   "DB_SDC_GLOBAL_EMS_ID_ACT" : Int = PLC DB_SDC_GLOBAL.EMS_ID_ACT AT %DB3700.DBW0, 1 s   // Aktuelle Anzahl der EMS-Treiber / Current quantity of EMS drivers
   "DB_SDC_GLOBAL_SYNCH[3].MAX_FAKT" : Real = PLC DB_SDC_GLOBAL.SYNCH[3].MAX_FAKT AT %DB3700.DBD214, 1 s   // Faktor für maximale Synchronisiergeschwindigkeit / Faktor Speed for Synchron MAX
   "DB_SDC_GLOBAL_SYNCH[13].SET_DIST" : Int = PLC DB_SDC_GLOBAL.SYNCH[13].SET_DIST AT %DB3700.DBW384, 1 s   // Set point value: distance (mm)
   "DB_SDC_GLOBAL_LIMITS[3].RAPID_SLOW" : Int = PLC DB_SDC_GLOBAL.LIMITS[3].RAPID_SLOW AT %DB3700.DBW518, 1 s   // Umstellung Begrenzung auf Abstand (mm), Einschränkung / Changeover limit of distance (mm), limitation
   "DB_SDC_GLOBAL_SYNCH[3].K" : Real = PLC DB_SDC_GLOBAL.SYNCH[3].K AT %DB3700.DBD210, 1 s   // erreichen von Synchron Faktor / gain for Synchron Faktor
   "DB_SDC_GLOBAL_SYNCH[13].SYNCH_DIST" : Int = PLC DB_SDC_GLOBAL.SYNCH[13].SYNCH_DIST AT %DB3700.DBW386, 1 s   // Start synchron distance value: distance (mm)
   "DB_SDC_GLOBAL_SYNCH[5].SYNCH_DIST" : Int = PLC DB_SDC_GLOBAL.SYNCH[5].SYNCH_DIST AT %DB3700.DBW242, 1 s   // Start synchron distance value: distance (mm)
   "DB_SDC_GLOBAL_SYNCH[6].HYST" : Int = PLC DB_SDC_GLOBAL.SYNCH[6].HYST AT %DB3700.DBW262, 1 s   // IO Hysterese
   "DB_SDC_GLOBAL_SYNCH[14].HYST" : Int = PLC DB_SDC_GLOBAL.SYNCH[14].HYST AT %DB3700.DBW406, 1 s   // IO Hysterese
   "DB_SDC_GLOBAL_START_COURSE" : DInt = PLC DB_SDC_GLOBAL.START_COURSE AT %DB3700.DBD14, 1 s   // Start Barcodevalue of Course
   "DB_SDC_GLOBAL_SYNCH[0].MAX_FAKT" : Real = PLC DB_SDC_GLOBAL.SYNCH[0].MAX_FAKT AT %DB3700.DBD160, 1 s   // Faktor für maximale Synchronisiergeschwindigkeit / Faktor Speed for Synchron MAX
   "DB_SDC_GLOBAL_SYNCH[2].SET_DIST" : Int = PLC DB_SDC_GLOBAL.SYNCH[2].SET_DIST AT %DB3700.DBW186, 1 s   // Set point value: distance (mm)
   "DB_SDC_GLOBAL_LIMITS[4].SLOW_SPEED_FAKT" : Real = PLC DB_SDC_GLOBAL.LIMITS[4].SLOW_SPEED_FAKT AT %DB3700.DBD526, 1 s   // Faktor Geschwindigkeit für langsame Drehzahl / Faktor Speed for Slow Speed
   "DB_SDC_GLOBAL_LIMITS[5].SLOW_SPEED_FAKT" : Real = PLC DB_SDC_GLOBAL.LIMITS[5].SLOW_SPEED_FAKT AT %DB3700.DBD532, 1 s   // Faktor Geschwindigkeit für langsame Drehzahl / Faktor Speed for Slow Speed
   "DB_SDC_GLOBAL_MIN_DIST_EMS[15]" : Int = PLC DB_SDC_GLOBAL.MIN_DIST_EMS[15] AT %DB3700.DBW130, 1 s   // minimum distance
   "DB_SDC_GLOBAL_SYNCH[12].MIN_FAKT" : Real = PLC DB_SDC_GLOBAL.SYNCH[12].MIN_FAKT AT %DB3700.DBD380, 1 s   // Faktor für minimale Synchronisiergeschwindigkeit / Faktor Speed for Synchron MIN
   "DB_SDC_GLOBAL_SYNCH[14].MAX_FAKT" : Real = PLC DB_SDC_GLOBAL.SYNCH[14].MAX_FAKT AT %DB3700.DBD412, 1 s   // Faktor für maximale Synchronisiergeschwindigkeit / Faktor Speed for Synchron MAX
   "DB_SDC_GLOBAL_SYNCH[10].MAX_FAKT" : Real = PLC DB_SDC_GLOBAL.SYNCH[10].MAX_FAKT AT %DB3700.DBD340, 1 s   // Faktor für maximale Synchronisiergeschwindigkeit / Faktor Speed for Synchron MAX
   "DB_SDC_GLOBAL_SYNCH[8].SYNCH_DIST" : Int = PLC DB_SDC_GLOBAL.SYNCH[8].SYNCH_DIST AT %DB3700.DBW296, 1 s   // Start synchron distance value: distance (mm)
   "DB_SDC_GLOBAL_max_barcode_mm" : DInt = PLC DB_SDC_GLOBAL.max_barcode_mm AT %DB3700.DBD10, 1 s   // Upper limit, bar code value
   "DB_SDC_GLOBAL_LIMITS[4].RAPID_SLOW" : Int = PLC DB_SDC_GLOBAL.LIMITS[4].RAPID_SLOW AT %DB3700.DBW524, 1 s   // Umstellung Begrenzung auf Abstand (mm), Einschränkung / Changeover limit of distance (mm), limitation
   "DB_SDC_GLOBAL_SYNCH[3].SET_DIST" : Int = PLC DB_SDC_GLOBAL.SYNCH[3].SET_DIST AT %DB3700.DBW204, 1 s   // Set point value: distance (mm)
   "DB_SDC_GLOBAL_SYNCH[10].HYST" : Int = PLC DB_SDC_GLOBAL.SYNCH[10].HYST AT %DB3700.DBW334, 1 s   // IO Hysterese
   "DB_SDC_GLOBAL_MIN_DIST_EMS[4]" : Int = PLC DB_SDC_GLOBAL.MIN_DIST_EMS[4] AT %DB3700.DBW108, 1 s   // minimum distance
   "DB_SDC_GLOBAL_SYNCH[7].SYNCH_DIST" : Int = PLC DB_SDC_GLOBAL.SYNCH[7].SYNCH_DIST AT %DB3700.DBW278, 1 s   // Start synchron distance value: distance (mm)
   "DB_SDC_GLOBAL_SYNCH[4].K" : Real = PLC DB_SDC_GLOBAL.SYNCH[4].K AT %DB3700.DBD228, 1 s   // erreichen von Synchron Faktor / gain for Synchron Faktor
   "DB_SDC_GLOBAL_SYNCH[0].SET_DIST" : Int = PLC DB_SDC_GLOBAL.SYNCH[0].SET_DIST AT %DB3700.DBW150, 1 s   // Set point value: distance (mm)
   "DB_SDC_GLOBAL_LIMITS[10].SLOW_SPEED_FAKT" : Real = PLC DB_SDC_GLOBAL.LIMITS[10].SLOW_SPEED_FAKT AT %DB3700.DBD562, 1 s   // Faktor Geschwindigkeit für langsame Drehzahl / Faktor Speed for Slow Speed
   "DB_SDC_GLOBAL_MIN_DIST_EMS[10]" : Int = PLC DB_SDC_GLOBAL.MIN_DIST_EMS[10] AT %DB3700.DBW120, 1 s   // minimum distance
   "DB_SDC_GLOBAL_SYNCH[15].MAX_FAKT" : Real = PLC DB_SDC_GLOBAL.SYNCH[15].MAX_FAKT AT %DB3700.DBD430, 1 s   // Faktor für maximale Synchronisiergeschwindigkeit / Faktor Speed for Synchron MAX
   "DB_SDC_GLOBAL_SYNCH[12].MAX_FAKT" : Real = PLC DB_SDC_GLOBAL.SYNCH[12].MAX_FAKT AT %DB3700.DBD376, 1 s   // Faktor für maximale Synchronisiergeschwindigkeit / Faktor Speed for Synchron MAX
   "DB_SDC_GLOBAL_LIMITS[8].SLOW_SPEED_FAKT" : Real = PLC DB_SDC_GLOBAL.LIMITS[8].SLOW_SPEED_FAKT AT %DB3700.DBD550, 1 s   // Faktor Geschwindigkeit für langsame Drehzahl / Faktor Speed for Slow Speed
   "DB_SDC_GLOBAL_LIMITS[9].RAPID_SLOW" : Int = PLC DB_SDC_GLOBAL.LIMITS[9].RAPID_SLOW AT %DB3700.DBW554, 1 s   // Umstellung Begrenzung auf Abstand (mm), Einschränkung / Changeover limit of distance (mm), limitation
   "DB_SDC_GLOBAL_SYNCH[3].HYST" : Int = PLC DB_SDC_GLOBAL.SYNCH[3].HYST AT %DB3700.DBW208, 1 s   // IO Hysterese
   "DB_SDC_GLOBAL_SEK_CYCLE_COUNTER" : Int = PLC DB_SDC_GLOBAL.SEK_CYCLE_COUNTER AT %DB3700.DBW28, 1 s
   "DB_SDC_GLOBAL_EMS_VCleaner_1" : Int = PLC DB_SDC_GLOBAL.EMS_VCleaner_1 AT %DB3700.DBW90, 1 s

HMI tags "DB_SDC_HMI"
   "DB_SDC_GLOBAL_M.SDC_ER_Reset(1)" : Bool = PLC DB_SDC_GLOBAL.M.SDC_ER_Reset AT %DB3700.DBX600.4, 1 s   // Fehler Reset / Fault Reset

HMI tags "VAT_DB_SDC_TS_REFERENCE"
   "DB_SDC_TS_REFERENCE_3_HEADER.MAX_NR_SEK" : Int = PLC DB_SDC_TS_REFERENCE_3.HEADER.MAX_NR_SEK AT %DB3782.DBW4, 1 s   // Höchste SEK Nummer im DB
   "DB_SDC_TS_REFERENCE_1_HEADER.MIN_NR_SEK" : Int = PLC DB_SDC_TS_REFERENCE_1.HEADER.MIN_NR_SEK AT %DB3780.DBW2, 1 s   // Niedrigste SEK Nummer im DB
   "SDC\DB_SDC_TS_REFERENCE\_TS_Ref_Byte_80" : DInt, internal
   "SDC\DB_SDC_TS_REFERENCE\DB_SDC_TS_REFERENCE_X.Reference[XXX].Hoist_offset_3" : Array [0..15] of Char AT %DB0.DBX0.0, 1 s   // definition Hub-Offset 3(mm)
   "DB_SDC_TS_REFERENCE_5_HEADER.MIN_NR_SEK" : Int = PLC DB_SDC_TS_REFERENCE_5.HEADER.MIN_NR_SEK AT %DB3784.DBW2, 1 s   // Niedrigste SEK Nummer im DB
   "DB_SDC_TS_REFERENCE_6_HEADER.DB_NR" : Int = PLC DB_SDC_TS_REFERENCE_6.HEADER.DB_NR AT %DB3785.DBW0, 1 s   // DB Nummer
   "DB_SDC_TS_REFERENCE_2_HEADER.DB_NR" : Int = PLC DB_SDC_TS_REFERENCE_2.HEADER.DB_NR AT %DB3781.DBW0, 1 s   // DB Nummer
   "SDC\DB_SDC_TS_REFERENCE\DB_SDC_TS_REFERENCE_X.Reference[XXX].Height" : Array [0..15] of Char AT %DB0.DBX0.0, 1 s   // definition Hubposition (mm)
   "DB_SDC_TS_REFERENCE_3_HEADER.DB_NR" : Int = PLC DB_SDC_TS_REFERENCE_3.HEADER.DB_NR AT %DB3782.DBW0, 1 s   // DB Nummer
   "DB_SDC_TS_REFERENCE_2_HEADER.MAX_NR_SEK" : Int = PLC DB_SDC_TS_REFERENCE_2.HEADER.MAX_NR_SEK AT %DB3781.DBW4, 1 s   // Höchste SEK Nummer im DB
   "SDC\DB_SDC_TS_REFERENCE\_TS_Ref_DB_Nr" : Int, internal
   "SDC\DB_SDC_TS_REFERENCE\DB_SDC_TS_REFERENCE_X.Reference[XXX].Sektion" : Array [0..15] of Char AT %DB0.DBX0.0, 1 s   // definition Sektion
   "DB_SDC_TS_REFERENCE_1_HEADER.MAX_NR_SEK" : Int = PLC DB_SDC_TS_REFERENCE_1.HEADER.MAX_NR_SEK AT %DB3780.DBW4, 1 s   // Höchste SEK Nummer im DB
   "SDC\DB_SDC_TS_REFERENCE\_TS_Ref_Byte_32" : DInt, internal
   "SDC\DB_SDC_TS_REFERENCE\_TS_Ref_Byte_64" : DInt, internal
   "DB_SDC_TS_REFERENCE_6_HEADER.MIN_NR_SEK" : Int = PLC DB_SDC_TS_REFERENCE_6.HEADER.MIN_NR_SEK AT %DB3785.DBW2, 1 s   // Niedrigste SEK Nummer im DB
   "SDC\DB_SDC_TS_REFERENCE\DB_SDC_TS_REFERENCE_X.Reference[XXX].Hoist_offset_4" : Array [0..15] of Char AT %DB0.DBX0.0, 1 s   // definition Hub-Offset 4 (mm)
   "DB_SDC_TS_REFERENCE_1_HEADER.DB_NR" : Int = PLC DB_SDC_TS_REFERENCE_1.HEADER.DB_NR AT %DB3780.DBW0, 1 s   // DB Nummer
   "SDC\DB_SDC_TS_REFERENCE\_TS_Ref_Byte_16" : DInt, internal
   "SDC\DB_SDC_TS_REFERENCE\_TS_Ref_Byte_00" : DInt, internal
   "SDC\DB_SDC_TS_REFERENCE\DB_SDC_TS_REFERENCE_X.Reference[XXX].Hoist_offset_1" : Array [0..15] of Char AT %DB0.DBX0.0, 1 s   // definition Hub-Offset 1 (mm)
   "SDC\DB_SDC_TS_REFERENCE\_TS_Ref_Byte_48" : DInt, internal
   "SDC\DB_SDC_TS_REFERENCE\_TS_Ref_Byte_96" : DInt, internal
   "DB_SDC_TS_REFERENCE_1_HEADER.START_DAT" : Int = PLC DB_SDC_TS_REFERENCE_1.HEADER.START_DAT AT %DB3780.DBW6, 1 s   // Startadresse der SEK im DB
   "DB_SDC_TS_REFERENCE_1_HEADER.LAENGE_SEK_DATA" : Int = PLC DB_SDC_TS_REFERENCE_1.HEADER.LAENGE_SEK_DATA AT %DB3780.DBW8, 1 s   // Länge SEK Data
   "SDC\DB_SDC_TS_REFERENCE\DB_SDC_TS_REFERENCE_X.Reference[XXX].Actionpoint_2" : Array [0..15] of Char AT %DB0.DBX0.0, 1 s   // definition Actionpoint 2
   "DB_SDC_TS_REFERENCE_4_HEADER.MIN_NR_SEK" : Int = PLC DB_SDC_TS_REFERENCE_4.HEADER.MIN_NR_SEK AT %DB3783.DBW2, 1 s   // Niedrigste SEK Nummer im DB
   "SDC\DB_SDC_TS_REFERENCE\DB_SDC_TS_REFERENCE_X.Reference[XXX].Actionpoint_1" : Array [0..15] of Char AT %DB0.DBX0.0, 1 s   // definition Actionpoint 1
   "DB_SDC_TS_REFERENCE_2_HEADER.MIN_NR_SEK" : Int = PLC DB_SDC_TS_REFERENCE_2.HEADER.MIN_NR_SEK AT %DB3781.DBW2, 1 s   // Niedrigste SEK Nummer im DB
   "DB_SDC_TS_REFERENCE_5_HEADER.DB_NR" : Int = PLC DB_SDC_TS_REFERENCE_5.HEADER.DB_NR AT %DB3784.DBW0, 1 s   // DB Nummer
   "SDC\DB_SDC_TS_REFERENCE\_TS_Ref_Byte_112" : DInt, internal
   "DB_SDC_TS_REFERENCE_5_HEADER.MAX_NR_SEK" : Int = PLC DB_SDC_TS_REFERENCE_5.HEADER.MAX_NR_SEK AT %DB3784.DBW4, 1 s   // Höchste SEK Nummer im DB
   "DB_SDC_TS_REFERENCE_4_HEADER.DB_NR" : Int = PLC DB_SDC_TS_REFERENCE_4.HEADER.DB_NR AT %DB3783.DBW0, 1 s   // DB Nummer
   "SDC\DB_SDC_TS_REFERENCE\_TS_Ref_Nr" : Int, internal
      on ChangeValue: "SDC_TS_REFERENCE"("SDC\_TS_Nr")
   "DB_SDC_TS_REFERENCE_3_HEADER.MIN_NR_SEK" : Int = PLC DB_SDC_TS_REFERENCE_3.HEADER.MIN_NR_SEK AT %DB3782.DBW2, 1 s   // Niedrigste SEK Nummer im DB
   "DB_SDC_TS_REFERENCE_4_HEADER.MAX_NR_SEK" : Int = PLC DB_SDC_TS_REFERENCE_4.HEADER.MAX_NR_SEK AT %DB3783.DBW4, 1 s   // Höchste SEK Nummer im DB
   "DB_SDC_TS_REFERENCE_6_HEADER.MAX_NR_SEK" : Int = PLC DB_SDC_TS_REFERENCE_6.HEADER.MAX_NR_SEK AT %DB3785.DBW4, 1 s   // Höchste SEK Nummer im DB
   "SDC\DB_SDC_TS_REFERENCE\DB_SDC_TS_REFERENCE_X.Reference[XXX].Hoist_offset_2" : Array [0..15] of Char AT %DB0.DBX0.0, 1 s   // definition Hub-Offset 2 (mm)

HMI tags "DB_SDC_POSITION_INSERTS"
   "DB_SDC_BARCODE_INSERTS_INSERT[19].COURSELOW" : DInt = PLC DB_SDC_BARCODE_INSERTS.INSERT[19].COURSELOW AT %DB3734.DBD364, 1 s   // lower position value Course Barocdevalue befor Insert
   "DB_SDC_BARCODE_INSERTS_INSERT[4].COURSEHIGH" : DInt = PLC DB_SDC_BARCODE_INSERTS.INSERT[4].COURSEHIGH AT %DB3734.DBD68, 1 s   // höhere Positionswert Course Barocde Wert nach Insert / higher position value Course Barocdevalue after Insert
   "DB_SDC_BARCODE_INSERTS_INSERT[15].INSERTHIGH" : DInt = PLC DB_SDC_BARCODE_INSERTS.INSERT[15].INSERTHIGH AT %DB3734.DBD296, 1 s   // höhere Positionswert Barocde Wert liegt Hoch / higher position value Barocdevalue Insert high
   "DB_SDC_BARCODE_INSERTS_INSERT[8].COURSELOW" : DInt = PLC DB_SDC_BARCODE_INSERTS.INSERT[8].COURSELOW AT %DB3734.DBD144, 1 s   // lower position value Course Barocdevalue befor Insert
   "DB_SDC_BARCODE_INSERTS_INSERT[9].INSERTLOW" : DInt = PLC DB_SDC_BARCODE_INSERTS.INSERT[9].INSERTLOW AT %DB3734.DBD172, 1 s   // lower position value Barocdevalue Insert low
   "DB_SDC_BARCODE_INSERTS_INSERT[14].COURSELOW" : DInt = PLC DB_SDC_BARCODE_INSERTS.INSERT[14].COURSELOW AT %DB3734.DBD264, 1 s   // lower position value Course Barocdevalue befor Insert
   "DB_SDC_BARCODE_INSERTS_INSERT[15].COURSEHIGH" : DInt = PLC DB_SDC_BARCODE_INSERTS.INSERT[15].COURSEHIGH AT %DB3734.DBD288, 1 s   // höhere Positionswert Course Barocde Wert nach Insert / higher position value Course Barocdevalue after Insert
   "DB_SDC_BARCODE_INSERTS_INSERT[19].COURSEHIGH" : DInt = PLC DB_SDC_BARCODE_INSERTS.INSERT[19].COURSEHIGH AT %DB3734.DBD368, 1 s   // höhere Positionswert Course Barocde Wert nach Insert / higher position value Course Barocdevalue after Insert
   "DB_SDC_BARCODE_INSERTS_INSERT[17].INSERTLOW" : DInt = PLC DB_SDC_BARCODE_INSERTS.INSERT[17].INSERTLOW AT %DB3734.DBD332, 1 s   // lower position value Barocdevalue Insert low
   "DB_SDC_BARCODE_INSERTS_INSERT[16].COURSEHIGH" : DInt = PLC DB_SDC_BARCODE_INSERTS.INSERT[16].COURSEHIGH AT %DB3734.DBD308, 1 s   // höhere Positionswert Course Barocde Wert nach Insert / higher position value Course Barocdevalue after Insert
   "DB_SDC_BARCODE_INSERTS_HYST" : Int = PLC DB_SDC_BARCODE_INSERTS.HYST AT %DB3734.DBW0, 1 s   // Hysterese für Positionswerte
   "DB_SDC_BARCODE_INSERTS_INSERT[3].OFFSET" : DInt = PLC DB_SDC_BARCODE_INSERTS.INSERT[3].OFFSET AT %DB3734.DBD60, 1 s   // absoluten Offset zu Beginn der Einfügen -> zusätzlich von allen Einsätzen unter / absolute offset at the start of the Insert -> addition from all inserts below
   "DB_SDC_BARCODE_INSERTS_INSERT[16].OFFSET" : DInt = PLC DB_SDC_BARCODE_INSERTS.INSERT[16].OFFSET AT %DB3734.DBD320, 1 s   // absoluten Offset zu Beginn der Einfügen -> zusätzlich von allen Einsätzen unter / absolute offset at the start of the Insert -> addition from all inserts below
   "DB_SDC_BARCODE_INSERTS_INSERT[10].OFFSET" : DInt = PLC DB_SDC_BARCODE_INSERTS.INSERT[10].OFFSET AT %DB3734.DBD200, 1 s   // absoluten Offset zu Beginn der Einfügen -> zusätzlich von allen Einsätzen unter / absolute offset at the start of the Insert -> addition from all inserts below
   "DB_SDC_BARCODE_INSERTS_INSERT[17].COURSELOW" : DInt = PLC DB_SDC_BARCODE_INSERTS.INSERT[17].COURSELOW AT %DB3734.DBD324, 1 s   // lower position value Course Barocdevalue befor Insert
   "DB_SDC_BARCODE_INSERTS_INSERT[4].INSERTLOW" : DInt = PLC DB_SDC_BARCODE_INSERTS.INSERT[4].INSERTLOW AT %DB3734.DBD72, 1 s   // lower position value Barocdevalue Insert low
   "DB_SDC_BARCODE_INSERTS_INSERT[20].COURSELOW" : DInt = PLC DB_SDC_BARCODE_INSERTS.INSERT[20].COURSELOW AT %DB3734.DBD384, 1 s   // lower position value Course Barocdevalue befor Insert
   "DB_SDC_BARCODE_INSERTS_INSERT[12].COURSELOW" : DInt = PLC DB_SDC_BARCODE_INSERTS.INSERT[12].COURSELOW AT %DB3734.DBD224, 1 s   // lower position value Course Barocdevalue befor Insert
   "DB_SDC_BARCODE_INSERTS_INSERT[7].COURSELOW" : DInt = PLC DB_SDC_BARCODE_INSERTS.INSERT[7].COURSELOW AT %DB3734.DBD124, 1 s   // lower position value Course Barocdevalue befor Insert
   "DB_SDC_BARCODE_INSERTS_INSERT[10].COURSELOW" : DInt = PLC DB_SDC_BARCODE_INSERTS.INSERT[10].COURSELOW AT %DB3734.DBD184, 1 s   // lower position value Course Barocdevalue befor Insert
   "DB_SDC_BARCODE_INSERTS_INSERT[3].COURSELOW" : DInt = PLC DB_SDC_BARCODE_INSERTS.INSERT[3].COURSELOW AT %DB3734.DBD44, 1 s   // lower position value Course Barocdevalue befor Insert
   "DB_SDC_BARCODE_INSERTS_INSERT[11].COURSELOW" : DInt = PLC DB_SDC_BARCODE_INSERTS.INSERT[11].COURSELOW AT %DB3734.DBD204, 1 s   // lower position value Course Barocdevalue befor Insert
   "DB_SDC_BARCODE_INSERTS_INSERT[15].COURSELOW" : DInt = PLC DB_SDC_BARCODE_INSERTS.INSERT[15].COURSELOW AT %DB3734.DBD284, 1 s   // lower position value Course Barocdevalue befor Insert
   "DB_SDC_BARCODE_INSERTS_INSERT[11].INSERTHIGH" : DInt = PLC DB_SDC_BARCODE_INSERTS.INSERT[11].INSERTHIGH AT %DB3734.DBD216, 1 s   // höhere Positionswert Barocde Wert liegt Hoch / higher position value Barocdevalue Insert high
   "DB_SDC_BARCODE_INSERTS_INSERT[17].INSERTHIGH" : DInt = PLC DB_SDC_BARCODE_INSERTS.INSERT[17].INSERTHIGH AT %DB3734.DBD336, 1 s   // höhere Positionswert Barocde Wert liegt Hoch / higher position value Barocdevalue Insert high
   "DB_SDC_BARCODE_INSERTS_INSERT[1].COURSEHIGH" : DInt = PLC DB_SDC_BARCODE_INSERTS.INSERT[1].COURSEHIGH AT %DB3734.DBD8, 1 s   // höhere Positionswert Course Barocde Wert nach Insert / higher position value Course Barocdevalue after Insert
   "DB_SDC_BARCODE_INSERTS_INSERT[11].OFFSET" : DInt = PLC DB_SDC_BARCODE_INSERTS.INSERT[11].OFFSET AT %DB3734.DBD220, 1 s   // absoluten Offset zu Beginn der Einfügen -> zusätzlich von allen Einsätzen unter / absolute offset at the start of the Insert -> addition from all inserts below
   "DB_SDC_BARCODE_INSERTS_INSERT[7].INSERTLOW" : DInt = PLC DB_SDC_BARCODE_INSERTS.INSERT[7].INSERTLOW AT %DB3734.DBD132, 1 s   // lower position value Barocdevalue Insert low
   "DB_SDC_BARCODE_INSERTS_INSERT[12].INSERTLOW" : DInt = PLC DB_SDC_BARCODE_INSERTS.INSERT[12].INSERTLOW AT %DB3734.DBD232, 1 s   // lower position value Barocdevalue Insert low
   "DB_SDC_BARCODE_INSERTS_INSERT[10].COURSEHIGH" : DInt = PLC DB_SDC_BARCODE_INSERTS.INSERT[10].COURSEHIGH AT %DB3734.DBD188, 1 s   // höhere Positionswert Course Barocde Wert nach Insert / higher position value Course Barocdevalue after Insert
   "DB_SDC_BARCODE_INSERTS_INSERTS" : Int = PLC DB_SDC_BARCODE_INSERTS.INSERTS AT %DB3734.DBW2, 1 s   // Positioning Leaps
   "DB_SDC_BARCODE_INSERTS_INSERT[8].INSERTHIGH" : DInt = PLC DB_SDC_BARCODE_INSERTS.INSERT[8].INSERTHIGH AT %DB3734.DBD156, 1 s   // höhere Positionswert Barocde Wert liegt Hoch / higher position value Barocdevalue Insert high
   "DB_SDC_BARCODE_INSERTS_INSERT[18].COURSELOW" : DInt = PLC DB_SDC_BARCODE_INSERTS.INSERT[18].COURSELOW AT %DB3734.DBD344, 1 s   // lower position value Course Barocdevalue befor Insert
   "DB_SDC_BARCODE_INSERTS_INSERT[5].INSERTHIGH" : DInt = PLC DB_SDC_BARCODE_INSERTS.INSERT[5].INSERTHIGH AT %DB3734.DBD96, 1 s   // höhere Positionswert Barocde Wert liegt Hoch / higher position value Barocdevalue Insert high
   "DB_SDC_BARCODE_INSERTS_INSERT[16].INSERTLOW" : DInt = PLC DB_SDC_BARCODE_INSERTS.INSERT[16].INSERTLOW AT %DB3734.DBD312, 1 s   // lower position value Barocdevalue Insert low
   "DB_SDC_BARCODE_INSERTS_INSERT[19].INSERTHIGH" : DInt = PLC DB_SDC_BARCODE_INSERTS.INSERT[19].INSERTHIGH AT %DB3734.DBD376, 1 s   // höhere Positionswert Barocde Wert liegt Hoch / higher position value Barocdevalue Insert high
   "DB_SDC_BARCODE_INSERTS_INSERT[18].COURSEHIGH" : DInt = PLC DB_SDC_BARCODE_INSERTS.INSERT[18].COURSEHIGH AT %DB3734.DBD348, 1 s   // höhere Positionswert Course Barocde Wert nach Insert / higher position value Course Barocdevalue after Insert
   "DB_SDC_BARCODE_INSERTS_INSERT[19].OFFSET" : DInt = PLC DB_SDC_BARCODE_INSERTS.INSERT[19].OFFSET AT %DB3734.DBD380, 1 s   // absoluten Offset zu Beginn der Einfügen -> zusätzlich von allen Einsätzen unter / absolute offset at the start of the Insert -> addition from all inserts below
   "DB_SDC_BARCODE_INSERTS_INSERT[8].INSERTLOW" : DInt = PLC DB_SDC_BARCODE_INSERTS.INSERT[8].INSERTLOW AT %DB3734.DBD152, 1 s   // lower position value Barocdevalue Insert low
   "DB_SDC_BARCODE_INSERTS_ABS_DIST_COURSE" : DInt = PLC DB_SDC_BARCODE_INSERTS.ABS_DIST_COURSE AT %DB3734.DBD404, 1 s   // abslolute Entfernung / abslolute Distance Course
   "DB_SDC_BARCODE_INSERTS_INSERT[14].INSERTLOW" : DInt = PLC DB_SDC_BARCODE_INSERTS.INSERT[14].INSERTLOW AT %DB3734.DBD272, 1 s   // lower position value Barocdevalue Insert low
   "DB_SDC_BARCODE_INSERTS_INSERT[13].COURSEHIGH" : DInt = PLC DB_SDC_BARCODE_INSERTS.INSERT[13].COURSEHIGH AT %DB3734.DBD248, 1 s   // höhere Positionswert Course Barocde Wert nach Insert / higher position value Course Barocdevalue after Insert
   "DB_SDC_BARCODE_INSERTS_INSERT[14].INSERTHIGH" : DInt = PLC DB_SDC_BARCODE_INSERTS.INSERT[14].INSERTHIGH AT %DB3734.DBD276, 1 s   // höhere Positionswert Barocde Wert liegt Hoch / higher position value Barocdevalue Insert high
   "DB_SDC_BARCODE_INSERTS_INSERT[5].INSERTLOW" : DInt = PLC DB_SDC_BARCODE_INSERTS.INSERT[5].INSERTLOW AT %DB3734.DBD92, 1 s   // lower position value Barocdevalue Insert low
   "DB_SDC_BARCODE_INSERTS_INSERT[14].OFFSET" : DInt = PLC DB_SDC_BARCODE_INSERTS.INSERT[14].OFFSET AT %DB3734.DBD280, 1 s   // absoluten Offset zu Beginn der Einfügen -> zusätzlich von allen Einsätzen unter / absolute offset at the start of the Insert -> addition from all inserts below
   "DB_SDC_BARCODE_INSERTS_INSERT[13].COURSELOW" : DInt = PLC DB_SDC_BARCODE_INSERTS.INSERT[13].COURSELOW AT %DB3734.DBD244, 1 s   // lower position value Course Barocdevalue befor Insert
   "DB_SDC_BARCODE_INSERTS_INSERT[7].COURSEHIGH" : DInt = PLC DB_SDC_BARCODE_INSERTS.INSERT[7].COURSEHIGH AT %DB3734.DBD128, 1 s   // höhere Positionswert Course Barocde Wert nach Insert / higher position value Course Barocdevalue after Insert
   "DB_SDC_BARCODE_INSERTS_INSERT[12].COURSEHIGH" : DInt = PLC DB_SDC_BARCODE_INSERTS.INSERT[12].COURSEHIGH AT %DB3734.DBD228, 1 s   // höhere Positionswert Course Barocde Wert nach Insert / higher position value Course Barocdevalue after Insert
   "DB_SDC_BARCODE_INSERTS_INSERT[18].INSERTHIGH" : DInt = PLC DB_SDC_BARCODE_INSERTS.INSERT[18].INSERTHIGH AT %DB3734.DBD356, 1 s   // höhere Positionswert Barocde Wert liegt Hoch / higher position value Barocdevalue Insert high
   "DB_SDC_BARCODE_INSERTS_INSERT[1].OFFSET" : DInt = PLC DB_SDC_BARCODE_INSERTS.INSERT[1].OFFSET AT %DB3734.DBD20, 1 s   // absoluten Offset zu Beginn der Einfügen -> zusätzlich von allen Einsätzen unter / absolute offset at the start of the Insert -> addition from all inserts below
   "DB_SDC_BARCODE_INSERTS_INSERT[1].INSERTHIGH" : DInt = PLC DB_SDC_BARCODE_INSERTS.INSERT[1].INSERTHIGH AT %DB3734.DBD16, 1 s   // höhere Positionswert Barocde Wert liegt Hoch / higher position value Barocdevalue Insert high
   "DB_SDC_BARCODE_INSERTS_INSERT[1].COURSELOW" : DInt = PLC DB_SDC_BARCODE_INSERTS.INSERT[1].COURSELOW AT %DB3734.DBD4, 1 s   // lower position value Course Barocdevalue befor Insert
   "DB_SDC_BARCODE_INSERTS_INSERT[3].INSERTHIGH" : DInt = PLC DB_SDC_BARCODE_INSERTS.INSERT[3].INSERTHIGH AT %DB3734.DBD56, 1 s   // höhere Positionswert Barocde Wert liegt Hoch / higher position value Barocdevalue Insert high
   "DB_SDC_BARCODE_INSERTS_INSERT[8].COURSEHIGH" : DInt = PLC DB_SDC_BARCODE_INSERTS.INSERT[8].COURSEHIGH AT %DB3734.DBD148, 1 s   // höhere Positionswert Course Barocde Wert nach Insert / higher position value Course Barocdevalue after Insert
   "DB_SDC_BARCODE_INSERTS_INSERT[5].OFFSET" : DInt = PLC DB_SDC_BARCODE_INSERTS.INSERT[5].OFFSET AT %DB3734.DBD100, 1 s   // absoluten Offset zu Beginn der Einfügen -> zusätzlich von allen Einsätzen unter / absolute offset at the start of the Insert -> addition from all inserts below
   "DB_SDC_BARCODE_INSERTS_INSERT[9].COURSELOW" : DInt = PLC DB_SDC_BARCODE_INSERTS.INSERT[9].COURSELOW AT %DB3734.DBD164, 1 s   // lower position value Course Barocdevalue befor Insert
   "DB_SDC_BARCODE_INSERTS_INSERT[14].COURSEHIGH" : DInt = PLC DB_SDC_BARCODE_INSERTS.INSERT[14].COURSEHIGH AT %DB3734.DBD268, 1 s   // höhere Positionswert Course Barocde Wert nach Insert / higher position value Course Barocdevalue after Insert
   "DB_SDC_BARCODE_INSERTS_INSERT[2].OFFSET" : DInt = PLC DB_SDC_BARCODE_INSERTS.INSERT[2].OFFSET AT %DB3734.DBD40, 1 s   // absoluten Offset zu Beginn der Einfügen -> zusätzlich von allen Einsätzen unter / absolute offset at the start of the Insert -> addition from all inserts below
   "DB_SDC_BARCODE_INSERTS_INSERT[17].OFFSET" : DInt = PLC DB_SDC_BARCODE_INSERTS.INSERT[17].OFFSET AT %DB3734.DBD340, 1 s   // absoluten Offset zu Beginn der Einfügen -> zusätzlich von allen Einsätzen unter / absolute offset at the start of the Insert -> addition from all inserts below
   "DB_SDC_BARCODE_INSERTS_INSERT[2].COURSELOW" : DInt = PLC DB_SDC_BARCODE_INSERTS.INSERT[2].COURSELOW AT %DB3734.DBD24, 1 s   // lower position value Course Barocdevalue befor Insert
   "DB_SDC_BARCODE_INSERTS_INSERT[16].COURSELOW" : DInt = PLC DB_SDC_BARCODE_INSERTS.INSERT[16].COURSELOW AT %DB3734.DBD304, 1 s   // lower position value Course Barocdevalue befor Insert
   "DB_SDC_BARCODE_INSERTS_INSERT[13].INSERTHIGH" : DInt = PLC DB_SDC_BARCODE_INSERTS.INSERT[13].INSERTHIGH AT %DB3734.DBD256, 1 s   // höhere Positionswert Barocde Wert liegt Hoch / higher position value Barocdevalue Insert high
   "DB_SDC_BARCODE_INSERTS_INSERT[2].INSERTHIGH" : DInt = PLC DB_SDC_BARCODE_INSERTS.INSERT[2].INSERTHIGH AT %DB3734.DBD36, 1 s   // höhere Positionswert Barocde Wert liegt Hoch / higher position value Barocdevalue Insert high
   "DB_SDC_BARCODE_INSERTS_INSERT[11].INSERTLOW" : DInt = PLC DB_SDC_BARCODE_INSERTS.INSERT[11].INSERTLOW AT %DB3734.DBD212, 1 s   // lower position value Barocdevalue Insert low
   "DB_SDC_BARCODE_INSERTS_INSERT[16].INSERTHIGH" : DInt = PLC DB_SDC_BARCODE_INSERTS.INSERT[16].INSERTHIGH AT %DB3734.DBD316, 1 s   // höhere Positionswert Barocde Wert liegt Hoch / higher position value Barocdevalue Insert high
   "DB_SDC_BARCODE_INSERTS_INSERT[20].COURSEHIGH" : DInt = PLC DB_SDC_BARCODE_INSERTS.INSERT[20].COURSEHIGH AT %DB3734.DBD388, 1 s   // höhere Positionswert Course Barocde Wert nach Insert / higher position value Course Barocdevalue after Insert
   "DB_SDC_BARCODE_INSERTS_INSERT[2].COURSEHIGH" : DInt = PLC DB_SDC_BARCODE_INSERTS.INSERT[2].COURSEHIGH AT %DB3734.DBD28, 1 s   // höhere Positionswert Course Barocde Wert nach Insert / higher position value Course Barocdevalue after Insert
   "DB_SDC_BARCODE_INSERTS_INSERT[5].COURSEHIGH" : DInt = PLC DB_SDC_BARCODE_INSERTS.INSERT[5].COURSEHIGH AT %DB3734.DBD88, 1 s   // höhere Positionswert Course Barocde Wert nach Insert / higher position value Course Barocdevalue after Insert
   "DB_SDC_BARCODE_INSERTS_INSERT[18].INSERTLOW" : DInt = PLC DB_SDC_BARCODE_INSERTS.INSERT[18].INSERTLOW AT %DB3734.DBD352, 1 s   // lower position value Barocdevalue Insert low
   "DB_SDC_BARCODE_INSERTS_INSERT[20].INSERTHIGH" : DInt = PLC DB_SDC_BARCODE_INSERTS.INSERT[20].INSERTHIGH AT %DB3734.DBD396, 1 s   // höhere Positionswert Barocde Wert liegt Hoch / higher position value Barocdevalue Insert high
   "DB_SDC_BARCODE_INSERTS_INSERT[15].OFFSET" : DInt = PLC DB_SDC_BARCODE_INSERTS.INSERT[15].OFFSET AT %DB3734.DBD300, 1 s   // absoluten Offset zu Beginn der Einfügen -> zusätzlich von allen Einsätzen unter / absolute offset at the start of the Insert -> addition from all inserts below
   "DB_SDC_BARCODE_INSERTS_INSERT[5].COURSELOW" : DInt = PLC DB_SDC_BARCODE_INSERTS.INSERT[5].COURSELOW AT %DB3734.DBD84, 1 s   // lower position value Course Barocdevalue befor Insert
   "DB_SDC_BARCODE_INSERTS_INSERT[2].INSERTLOW" : DInt = PLC DB_SDC_BARCODE_INSERTS.INSERT[2].INSERTLOW AT %DB3734.DBD32, 1 s   // lower position value Barocdevalue Insert low
   "DB_SDC_BARCODE_INSERTS_INSERT[12].OFFSET" : DInt = PLC DB_SDC_BARCODE_INSERTS.INSERT[12].OFFSET AT %DB3734.DBD240, 1 s   // absoluten Offset zu Beginn der Einfügen -> zusätzlich von allen Einsätzen unter / absolute offset at the start of the Insert -> addition from all inserts below
   "DB_SDC_BARCODE_INSERTS_INSERT[17].COURSEHIGH" : DInt = PLC DB_SDC_BARCODE_INSERTS.INSERT[17].COURSEHIGH AT %DB3734.DBD328, 1 s   // höhere Positionswert Course Barocde Wert nach Insert / higher position value Course Barocdevalue after Insert
   "DB_SDC_BARCODE_INSERTS_INSERT[4].INSERTHIGH" : DInt = PLC DB_SDC_BARCODE_INSERTS.INSERT[4].INSERTHIGH AT %DB3734.DBD76, 1 s   // höhere Positionswert Barocde Wert liegt Hoch / higher position value Barocdevalue Insert high
   "DB_SDC_BARCODE_INSERTS_INSERT[20].INSERTLOW" : DInt = PLC DB_SDC_BARCODE_INSERTS.INSERT[20].INSERTLOW AT %DB3734.DBD392, 1 s   // lower position value Barocdevalue Insert low
   "DB_SDC_BARCODE_INSERTS_INSERT[10].INSERTLOW" : DInt = PLC DB_SDC_BARCODE_INSERTS.INSERT[10].INSERTLOW AT %DB3734.DBD192, 1 s   // lower position value Barocdevalue Insert low
   "DB_SDC_BARCODE_INSERTS_INSERT[20].OFFSET" : DInt = PLC DB_SDC_BARCODE_INSERTS.INSERT[20].OFFSET AT %DB3734.DBD400, 1 s   // absoluten Offset zu Beginn der Einfügen -> zusätzlich von allen Einsätzen unter / absolute offset at the start of the Insert -> addition from all inserts below
   "DB_SDC_BARCODE_INSERTS_INSERT[4].COURSELOW" : DInt = PLC DB_SDC_BARCODE_INSERTS.INSERT[4].COURSELOW AT %DB3734.DBD64, 1 s   // lower position value Course Barocdevalue befor Insert
   "DB_SDC_BARCODE_INSERTS_INSERT[3].COURSEHIGH" : DInt = PLC DB_SDC_BARCODE_INSERTS.INSERT[3].COURSEHIGH AT %DB3734.DBD48, 1 s   // höhere Positionswert Course Barocde Wert nach Insert / higher position value Course Barocdevalue after Insert
   "DB_SDC_BARCODE_INSERTS_INSERT[6].COURSELOW" : DInt = PLC DB_SDC_BARCODE_INSERTS.INSERT[6].COURSELOW AT %DB3734.DBD104, 1 s   // lower position value Course Barocdevalue befor Insert
   "DB_SDC_BARCODE_INSERTS_INSERT[6].COURSEHIGH" : DInt = PLC DB_SDC_BARCODE_INSERTS.INSERT[6].COURSEHIGH AT %DB3734.DBD108, 1 s   // höhere Positionswert Course Barocde Wert nach Insert / higher position value Course Barocdevalue after Insert
   "DB_SDC_BARCODE_INSERTS_INSERT[3].INSERTLOW" : DInt = PLC DB_SDC_BARCODE_INSERTS.INSERT[3].INSERTLOW AT %DB3734.DBD52, 1 s   // lower position value Barocdevalue Insert low
   "DB_SDC_BARCODE_INSERTS_INSERT[12].INSERTHIGH" : DInt = PLC DB_SDC_BARCODE_INSERTS.INSERT[12].INSERTHIGH AT %DB3734.DBD236, 1 s   // höhere Positionswert Barocde Wert liegt Hoch / higher position value Barocdevalue Insert high
   "DB_SDC_BARCODE_INSERTS_INSERT[9].OFFSET" : DInt = PLC DB_SDC_BARCODE_INSERTS.INSERT[9].OFFSET AT %DB3734.DBD180, 1 s   // absoluten Offset zu Beginn der Einfügen -> zusätzlich von allen Einsätzen unter / absolute offset at the start of the Insert -> addition from all inserts below
   "DB_SDC_BARCODE_INSERTS_INSERT[9].COURSEHIGH" : DInt = PLC DB_SDC_BARCODE_INSERTS.INSERT[9].COURSEHIGH AT %DB3734.DBD168, 1 s   // höhere Positionswert Course Barocde Wert nach Insert / higher position value Course Barocdevalue after Insert
   "DB_SDC_BARCODE_INSERTS_INSERT[6].INSERTHIGH" : DInt = PLC DB_SDC_BARCODE_INSERTS.INSERT[6].INSERTHIGH AT %DB3734.DBD116, 1 s   // höhere Positionswert Barocde Wert liegt Hoch / higher position value Barocdevalue Insert high
   "DB_SDC_BARCODE_INSERTS_INSERT[6].INSERTLOW" : DInt = PLC DB_SDC_BARCODE_INSERTS.INSERT[6].INSERTLOW AT %DB3734.DBD112, 1 s   // lower position value Barocdevalue Insert low
   "DB_SDC_BARCODE_INSERTS_INSERT[7].INSERTHIGH" : DInt = PLC DB_SDC_BARCODE_INSERTS.INSERT[7].INSERTHIGH AT %DB3734.DBD136, 1 s   // höhere Positionswert Barocde Wert liegt Hoch / higher position value Barocdevalue Insert high
   "DB_SDC_BARCODE_INSERTS_INSERT[15].INSERTLOW" : DInt = PLC DB_SDC_BARCODE_INSERTS.INSERT[15].INSERTLOW AT %DB3734.DBD292, 1 s   // lower position value Barocdevalue Insert low
   "DB_SDC_BARCODE_INSERTS_INSERT[4].OFFSET" : DInt = PLC DB_SDC_BARCODE_INSERTS.INSERT[4].OFFSET AT %DB3734.DBD80, 1 s   // absoluten Offset zu Beginn der Einfügen -> zusätzlich von allen Einsätzen unter / absolute offset at the start of the Insert -> addition from all inserts below
   "DB_SDC_BARCODE_INSERTS_INSERT[9].INSERTHIGH" : DInt = PLC DB_SDC_BARCODE_INSERTS.INSERT[9].INSERTHIGH AT %DB3734.DBD176, 1 s   // höhere Positionswert Barocde Wert liegt Hoch / higher position value Barocdevalue Insert high
   "DB_SDC_BARCODE_INSERTS_INSERT[6].OFFSET" : DInt = PLC DB_SDC_BARCODE_INSERTS.INSERT[6].OFFSET AT %DB3734.DBD120, 1 s   // absoluten Offset zu Beginn der Einfügen -> zusätzlich von allen Einsätzen unter / absolute offset at the start of the Insert -> addition from all inserts below
   "DB_SDC_BARCODE_INSERTS_INSERT[13].INSERTLOW" : DInt = PLC DB_SDC_BARCODE_INSERTS.INSERT[13].INSERTLOW AT %DB3734.DBD252, 1 s   // lower position value Barocdevalue Insert low
   "DB_SDC_BARCODE_INSERTS_INSERT[19].INSERTLOW" : DInt = PLC DB_SDC_BARCODE_INSERTS.INSERT[19].INSERTLOW AT %DB3734.DBD372, 1 s   // lower position value Barocdevalue Insert low
   "DB_SDC_BARCODE_INSERTS_INSERT[11].COURSEHIGH" : DInt = PLC DB_SDC_BARCODE_INSERTS.INSERT[11].COURSEHIGH AT %DB3734.DBD208, 1 s   // höhere Positionswert Course Barocde Wert nach Insert / higher position value Course Barocdevalue after Insert
   "DB_SDC_BARCODE_INSERTS_INSERT[8].OFFSET" : DInt = PLC DB_SDC_BARCODE_INSERTS.INSERT[8].OFFSET AT %DB3734.DBD160, 1 s   // absoluten Offset zu Beginn der Einfügen -> zusätzlich von allen Einsätzen unter / absolute offset at the start of the Insert -> addition from all inserts below
   "DB_SDC_BARCODE_INSERTS_INSERT[13].OFFSET" : DInt = PLC DB_SDC_BARCODE_INSERTS.INSERT[13].OFFSET AT %DB3734.DBD260, 1 s   // absoluten Offset zu Beginn der Einfügen -> zusätzlich von allen Einsätzen unter / absolute offset at the start of the Insert -> addition from all inserts below
   "DB_SDC_BARCODE_INSERTS_INSERT[7].OFFSET" : DInt = PLC DB_SDC_BARCODE_INSERTS.INSERT[7].OFFSET AT %DB3734.DBD140, 1 s   // absoluten Offset zu Beginn der Einfügen -> zusätzlich von allen Einsätzen unter / absolute offset at the start of the Insert -> addition from all inserts below
   "DB_SDC_BARCODE_INSERTS_INSERT[10].INSERTHIGH" : DInt = PLC DB_SDC_BARCODE_INSERTS.INSERT[10].INSERTHIGH AT %DB3734.DBD196, 1 s   // höhere Positionswert Barocde Wert liegt Hoch / higher position value Barocdevalue Insert high
   "DB_SDC_BARCODE_INSERTS_INSERT[1].INSERTLOW" : DInt = PLC DB_SDC_BARCODE_INSERTS.INSERT[1].INSERTLOW AT %DB3734.DBD12, 1 s   // lower position value Barocdevalue Insert low
   "DB_SDC_BARCODE_INSERTS_INSERT[18].OFFSET" : DInt = PLC DB_SDC_BARCODE_INSERTS.INSERT[18].OFFSET AT %DB3734.DBD360, 1 s   // absoluten Offset zu Beginn der Einfügen -> zusätzlich von allen Einsätzen unter / absolute offset at the start of the Insert -> addition from all inserts below

HMI tags "DB_SDC_EMS_INFO"
   "EMS_Zone[1]" : UDT_ZoneStructure = PLC EMS.Zone[1] AT %DB8.DBX1034.0, 1 s
   "EMS_Zone[2]" : UDT_ZoneStructure = PLC EMS.Zone[2] AT %DB8.DBX2068.0, 1 s
   "EMS_Zone[3]" : UDT_ZoneStructure = PLC EMS.Zone[3] AT %DB8.DBX3102.0, 1 s
   "EMS_Zone[7]" : UDT_ZoneStructure = PLC EMS.Zone[7] AT %DB8.DBX7238.0, 1 s
   "EMS_Zone[8]" : UDT_ZoneStructure = PLC EMS.Zone[8] AT %DB8.DBX8272.0, 1 s
   "EMS_Zone[9]" : UDT_ZoneStructure = PLC EMS.Zone[9] AT %DB8.DBX9306.0, 1 s
   "EMS_Zone[10]" : UDT_ZoneStructure = PLC EMS.Zone[10] AT %DB8.DBX10340.0, 1 s
   "EMS_Zone[11]" : UDT_ZoneStructure = PLC EMS.Zone[11] AT %DB8.DBX11374.0, 1 s
   "EMS_Zone[12]" : UDT_ZoneStructure = PLC EMS.Zone[12] AT %DB8.DBX12408.0, 1 s
   "EMS_Zone[13]" : UDT_ZoneStructure = PLC EMS.Zone[13] AT %DB8.DBX13442.0, 1 s
   "EMS_Zone[14]" : UDT_ZoneStructure = PLC EMS.Zone[14] AT %DB8.DBX14476.0, 1 s
   "EMS_Zone[15]" : UDT_ZoneStructure = PLC EMS.Zone[15] AT %DB8.DBX15510.0, 1 s
   "EMS_Zone[16]" : UDT_ZoneStructure = PLC EMS.Zone[16] AT %DB8.DBX16544.0, 1 s
   "EMS_Zone[17]" : UDT_ZoneStructure = PLC EMS.Zone[17] AT %DB8.DBX17578.0, 1 s
   "EMS_Zone[18]" : UDT_ZoneStructure = PLC EMS.Zone[18] AT %DB8.DBX18612.0, 1 s
   "EMS_Zone[19]" : UDT_ZoneStructure = PLC EMS.Zone[19] AT %DB8.DBX19646.0, 1 s
   "EMS_Zone[20]" : UDT_ZoneStructure = PLC EMS.Zone[20] AT %DB8.DBX20680.0, 1 s
   "EMS_Zone[21]" : UDT_ZoneStructure = PLC EMS.Zone[21] AT %DB8.DBX21714.0, 1 s
   "EMS_Zone[22]" : UDT_ZoneStructure = PLC EMS.Zone[22] AT %DB8.DBX22748.0, 1 s
   "EMS_Zone[23]" : UDT_ZoneStructure = PLC EMS.Zone[23] AT %DB8.DBX23782.0, 1 s
   "EMS_Zone[24]" : UDT_ZoneStructure = PLC EMS.Zone[24] AT %DB8.DBX24816.0, 1 s
   "EMS_Zone[25]" : UDT_ZoneStructure = PLC EMS.Zone[25] AT %DB8.DBX25850.0, 1 s
   "EMS_Zone[26]" : UDT_ZoneStructure = PLC EMS.Zone[26] AT %DB8.DBX26884.0, 1 s
   "EMS_Zone[27]" : UDT_ZoneStructure = PLC EMS.Zone[27] AT %DB8.DBX27918.0, 1 s
   "EMS_Zone[28]" : UDT_ZoneStructure = PLC EMS.Zone[28] AT %DB8.DBX28952.0, 1 s
   "EMS_Zone[29]" : UDT_ZoneStructure = PLC EMS.Zone[29] AT %DB8.DBX29986.0, 1 s
   "EMS_Zone[30]" : UDT_ZoneStructure = PLC EMS.Zone[30] AT %DB8.DBX31020.0, 1 s
   "EMS_Carrier[1]" : UDT_CarrierStructure = PLC EMS.Carrier[1] AT %DB8.DBX63156.0, 1 s
   "EMS_Carrier[2]" : UDT_CarrierStructure = PLC EMS.Carrier[2] AT %DB8.DBX63238.0, 1 s
   "EMS_Carrier[3]" : UDT_CarrierStructure = PLC EMS.Carrier[3] AT %DB8.DBX63320.0, 1 s
   "EMS_Carrier[4]" : UDT_CarrierStructure = PLC EMS.Carrier[4] AT %DB8.DBX63402.0, 1 s
   "EMS_Carrier[5]" : UDT_CarrierStructure = PLC EMS.Carrier[5] AT %DB8.DBX63484.0, 1 s
   "EMS_Carrier[6]" : UDT_CarrierStructure = PLC EMS.Carrier[6] AT %DB8.DBX63566.0, 1 s
   "EMS_Carrier[7]" : UDT_CarrierStructure = PLC EMS.Carrier[7] AT %DB8.DBX63648.0, 1 s
   "EMS_Carrier[8]" : UDT_CarrierStructure = PLC EMS.Carrier[8] AT %DB8.DBX63730.0, 1 s
   "EMS_Carrier[9]" : UDT_CarrierStructure = PLC EMS.Carrier[9] AT %DB8.DBX63812.0, 1 s
   "EMS_Carrier[10]" : UDT_CarrierStructure = PLC DB_SDC_ERRORS_STAT.ER_AKT[42].ER_STAT[3].DRIVE_POS AT %DB8.DBX63894.0, 1 s
   "EMS_Carrier[11]" : UDT_CarrierStructure = PLC EMS.Carrier[11] AT %DB8.DBX63976.0, 1 s
   "EMS_Carrier[12]" : UDT_CarrierStructure = PLC EMS.Carrier[12] AT %DB8.DBX64058.0, 1 s
   "EMS_Carrier[13]" : UDT_CarrierStructure = PLC EMS.Carrier[13] AT %DB8.DBX64140.0, 1 s
   "EMS_Carrier[14]" : UDT_CarrierStructure = PLC EMS.Carrier[14] AT %DB8.DBX64222.0, 1 s
   "EMS_Carrier[15]" : UDT_CarrierStructure = PLC EMS.Carrier[15] AT %DB8.DBX64304.0, 1 s
   "EMS_Carrier[16]" : UDT_CarrierStructure = PLC EMS.Carrier[16] AT %DB8.DBX64386.0, 1 s
   "EMS_Carrier[17]" : UDT_CarrierStructure = PLC EMS.Carrier[17] AT %DB8.DBX64468.0, 1 s
   "EMS_Carrier[18]" : UDT_CarrierStructure = PLC EMS.Carrier[18] AT %DB8.DBX64550.0, 1 s
   "EMS_Carrier[19]" : UDT_CarrierStructure = PLC EMS.Carrier[19] AT %DB8.DBX64632.0, 1 s
   "EMS_Carrier[20]" : UDT_CarrierStructure = PLC EMS.Carrier[20] AT %DB8.DBX64714.0, 1 s
   "EMS_Carrier[21]" : UDT_CarrierStructure = PLC EMS.Carrier[21] AT %DB8.DBX64796.0, 1 s
   "EMS_Carrier[22]" : UDT_CarrierStructure = PLC EMS.Carrier[22] AT %DB8.DBX64878.0, 1 s
   "EMS_Carrier[23]" : UDT_CarrierStructure = PLC EMS.Carrier[23] AT %DB8.DBX64960.0, 1 s
   "EMS_Carrier[24]" : UDT_CarrierStructure = PLC EMS.Carrier[24] AT %DB8.DBX65042.0, 1 s
   "EMS_Carrier[25]" : UDT_CarrierStructure = PLC EMS.Carrier[25] AT %DB8.DBX65124.0, 1 s
   "EMS_Carrier[26]" : UDT_CarrierStructure = PLC EMS.Carrier[26] AT %DB8.DBX65206.0, 1 s
   "EMS_Carrier[27]" : UDT_CarrierStructure = PLC EMS.Carrier[27] AT %DB8.DBX65288.0, 1 s
   "EMS_Carrier[28]" : UDT_CarrierStructure = PLC EMS.Carrier[28] AT %DB8.DBX65370.0, 1 s
   "EMS_Carrier[29]" : UDT_CarrierStructure = PLC EMS.Carrier[29] AT %DB8.DBX65452.0, 1 s
   "EMS_Carrier[30]" : UDT_CarrierStructure = PLC EMS.Carrier[30], 1 s
   "EMS_Carrier[31]" : UDT_CarrierStructure = PLC EMS.Carrier[31], 1 s
   "EMS_Carrier[32]" : UDT_CarrierStructure = PLC EMS.Carrier[32], 1 s
   "EMS_Carrier[33]" : UDT_CarrierStructure = PLC EMS.Carrier[33], 1 s
   "EMS_Carrier[34]" : UDT_CarrierStructure = PLC EMS.Carrier[34], 1 s
   "EMS_Carrier[35]" : UDT_CarrierStructure = PLC EMS.Carrier[35], 1 s
   "EMS_Carrier[36]" : UDT_CarrierStructure = PLC EMS.Carrier[36], 1 s
   "EMS_Carrier[37]" : UDT_CarrierStructure = PLC EMS.Carrier[37], 1 s
   "EMS_Carrier[38]" : UDT_CarrierStructure = PLC EMS.Carrier[38], 1 s
   "EMS_Carrier[39]" : UDT_CarrierStructure = PLC EMS.Carrier[39], 1 s
   "EMS_Carrier[40]" : UDT_CarrierStructure = PLC EMS.Carrier[40], 1 s

